// TIA Portal project "Energy_Drink_V15.1" (V15.1)

(* hardware
DEVICE "S7300/ET200M station_1"  S7-300 station
   slot 0: "Rail_0"  Rail  6ES7 390-1***0-0AA0
   slot 2: "ENERGY_DRINK_PROC"  CPU 314C-2 PN/DP  6ES7 314-6EH04-0AB0  V3.3
      slot 2: "PROFINET interface_1"  PN-IO
         slot 1: "Port_1"  Port
         slot 2: "Port_2"  Port
      slot 5: "DI 24/DO 16_1"  DI24/DO16
      slot 6: "AI 5/AO 2_1"  AI5/AO2
      slot 7: "Count_1"  Counter
      slot 8: "Positioning_1"  Positioning
   slot 4: "DI 16/DO 16x24VDC/0.5A_1"  DI16/DO16 x 24V / 0.5A  6ES7 323-1BL00-0AA0
   slot 5: "DI 8/DO 8x24VDC/0.5A_1"  DI8/DO8 x 24VDC / 0.5A  6ES7 323-1BH01-0AA0
   slot 6: "AI 2x12BIT_1"  AI2 x 12 bits  6ES7 331-7KB02-0AB0
   slot 7: "AO 4x12BIT_1"  AO4 x 12 bits  6ES7 332-5HD01-0AB0
DEVICE "HMI_1"  TP2200 Comfort
   slot 0: "HMI"  HMI  6AV2 124-0XC02-0AX0  13.0.1.0
   slot 1: "HMI_RT_1"  TP2200 Comfort  6AV2 124-0XC02-0AX0  13.0.1.0
   slot 5: "HMI_1.IE_CP_1"  Interfaz PROFINET
      slot 1: "Interfaz PROFINET_1"  Interfaz PROFINET
         slot 1: "Port_1"  Port
         slot 2: "Port_2"  Port
   slot 6: "HMI_1.IE_CP_2"  Interfaz PROFINET
      slot 1: "Interfaz PROFINET_GBit"  Interfaz PROFINET
         slot 1: "Port_1"  Port
   slot 7: "HMI_1.MPI/DP_CP_1"  Interfaz MPI/DP
*)

// ===== PLC "ENERGY_DRINK_PROC"  CPU 314C-2 PN/DP =====

VAR_GLOBAL   // PLC tag table "Default tag table"
   "M_Product_1" AT %MD100 : Real;
   "Tag_5" AT %MD50 : DWord;
   "Tag_6" AT %EW50 : Word;
   "Recipe_Num" AT %MW50 : Word;
   "M_Water_Flow" AT %MD112 : Real;
   "Num_Bach" AT %MW52 : Word;
   "Tag_3" AT %M10.0 : Bool;
   "Tag_7" AT %MD120 : Real;
   "Tag_13" AT %MD140 : Real;
   "M_Product_2" AT %MD104 : Real;
   "M_Product_3" AT %MD108 : Real;
   "M_Sirupe_Flow" AT %MD116 : Real;
   "FP_Conveyor_Act" AT %M255.7 : Bool;
   "FN_Bach_in_Prog" AT %M255.6 : Bool;
   "FN_TIMER.Q" AT %M255.5 : Bool;
   "FN_STOP_CMD" AT %M255.4 : Bool;
   "Tag_4" AT %MD200 : DWord;
   "Tag_10" AT %MW70 : Word;
   "Tag_11" AT %MD204 : DWord;
   "Tag_12" AT %M250.0 : Bool;
   "Tag_14" AT %M250.1 : Bool;
   "Tag_15" AT %MW60 : Int;
   "Tag_16" AT %MW62 : Int;
   "Tag_17" AT %MW64 : Int;
   "Tag_18" AT %MW66 : Int;
   "Tag_19" AT %MW68 : Int;
   "Tag_20" AT %MW72 : Int;
   "Tag_21" AT %MW74 : Int;
   "Tag_22" AT %MW76 : Int;
   "Tag_23" AT %MW78 : Int;
   "Tag_24" AT %MW80 : Int;
   "Tank1_Vlv" AT %AW800 : Word;
   "Tank2_Vlv" AT %AW802 : Word;
   "Tank3_Vlv" AT %AW804 : Word;
   "Sirupe_Vlv" AT %AW806 : Word;
   "Water_Vlv" AT %AW808 : Word;
   "Motor_VF" AT %AW810 : Word;
   "Tag_1" AT %MW82 : Int;
   "Tag_2" AT %M255.3 : Bool;
   "Tag_8" AT %M255.2 : Bool;
   "Tag_9" AT %M255.1 : Bool;
   "Tag_25" AT %M254.7 : Bool;
   "Tag_26" AT %M254.6 : Bool;
   "Tag_27" AT %M254.5 : Bool;
   "Total_Weight" AT %MD150 : Real;
   "Temp_Lim_Kg" AT %MD154 : Real;
   "Tag_29" AT %MD158 : Real;
   "Tag_28" AT %MD84 : DInt;
   "Tag_30" AT %M0.6 : Bool;
   "Tag_31" AT %M254.4 : Bool;
   "Tag_32" AT %M0.4 : Bool;
   "Tag_33" AT %M0.2 : Bool;
   "Tag_34" AT %M0.0 : Bool;
   "Tag_35" AT %M0.1 : Bool;
END_VAR

VAR_GLOBAL   // PLC tag table "VAR"
   "AUTO/MAN" AT %E0.0 : Bool;   // Switch Auto/Man
   "Start_Button" AT %E0.1 : Bool;   // Start switch "NO"
   "Stop_Button" AT %E0.2 : Bool;   // Stop switch "NC"
   "Emergency_Stop" AT %E0.3 : Bool;   // Emergency Stop "NC"
   "Man_Dis_Tk1_Vlv" AT %E136.1 : Bool;   // K1_Outlet gate Tank1 Switch
   "Man_Dis_Tk2_Vlv" AT %E136.2 : Bool;   // K2_Outlet gate Tank2 Switch
   "Man_Dis_Tk3_Vlv" AT %E136.3 : Bool;   // K3_Outlet gate Tank3 Switch
   "Man_Dis_Scale_Vlv" AT %E136.4 : Bool;   // K4_Outlet gate Scale Tank Switch
   "Convey_Man_Starter" AT %E136.5 : Bool;   // Starter start-delta motor Switch
   "Mixer_Man_Start" AT %E136.7 : Bool;   // VF Agitator motor Switch
   "Man_Dis_Mixer_Vlv" AT %E137.1 : Bool;   // K5_Outlet gate Mixer Tank Switch
   "Man_Water_Vlv" AT %E137.2 : Bool;   // K6_Water valve Switch
   "Man_Sirupe_Vlv" AT %E137.3 : Bool;   // K7_Sirupe valve Switch
   "Man_Fill_Tk1_Vlv" AT %E137.4 : Bool;   // K8_Filling valve Tank 1 Switch
   "Man_Fill_Tk2_Vlv" AT %E137.5 : Bool;   // K9_Filling valve Tank 2 Switch
   "Man_Fill_Tk3_Vlv" AT %E137.6 : Bool;   // K10_Filling valve Tank 3 Switch
   "OVL_Conveyor" AT %E137.7 : Bool;   // Overload Conveyor Motor
   "OVL_Mixer" AT %E138.0 : Bool;   // Overload VF Agitator
   "Recipe_1" AT %E138.1 : Bool;   // Recipe 1 Switch
   "Recipe_2" AT %E138.2 : Bool;   // Recipe 2 Switch
   "Recipe_3" AT %E138.3 : Bool;   // Recipe 3 Switch
   "Tank_1_Level" AT %EW800 : Int;
   "Tank_2_Level" AT %EW802 : Int;
   "Tank_3_Level" AT %EW804 : Int;
   "Weighing" AT %EW806 : Int;
   "Mixer_Tank_level" AT %EW808 : Int;
   "Water_Flow" AT %EW256 : Int;
   "Sirupe_Flow" AT %EW258 : Int;
   "Filling_Vlv_1_Opened" AT %E0.5 : Bool;
   "Filling_Vlv_1_Closed" AT %E0.6 : Bool;
   "Filling_Vlv_2_Closed" AT %E1.1 : Bool;
   "Filling_Vlv_2_Opened" AT %E1.2 : Bool;
   "Filling_Vlv_3_Closed" AT %E1.5 : Bool;
   "Filling_Vlv_3_Opened" AT %E1.6 : Bool;
   "Disch_Vlv_3_Opened" AT %E1.7 : Bool;
   "Disch_Vlv_3_Closed" AT %E2.0 : Bool;
   "Disch_Vlv_M_Opened" AT %E2.1 : Bool;
   "Disch_Vlv_M_Closed" AT %E2.2 : Bool;
   "Sirupe_Vlv_Closed" AT %E2.6 : Bool;
   "Disch_Vlv_1_Opened" AT %E0.7 : Bool;
   "Disch_Vlv_1_Closed" AT %E1.0 : Bool;
   "Disch_Vlv_2_Opened" AT %E1.3 : Bool;
   "Disch_Vlv_2_Closed" AT %E1.4 : Bool;
   "Water_Vlv_Closed" AT %E2.4 : Bool;
   "Water_Vlv_Opened" AT %E2.3 : Bool;
   "Sirupe_Vlv_Opened" AT %E2.5 : Bool;
   "Scale_Vlv_Opened" AT %E2.7 : Bool;
   "Scale_Vlv_Closed" AT %E136.0 : Bool;
   "Discharge_Vlv1" AT %A136.0 : Bool;   // Outlet gate Tank 1 rely
   "Discharge_Vlv2" AT %A136.1 : Bool;   // Outlet gate Tank 2 rely
   "Discharge_Vlv3" AT %A136.2 : Bool;   // Outlet gate Tank 3 rely
   "Scale_Dis_Vlv" AT %A136.3 : Bool;   // Outlet gate Scale Tank rely
   "Mixer_Dis_Vlv" AT %A136.4 : Bool;   // Outlet gate Mixer Tank rely
   "Filling_Vlv1" AT %A136.5 : Bool;   // Filling valve Tank 1 rely
   "Filling_Vlv2" AT %A136.6 : Bool;   // Filling valve Tank 2 rely
   "Filling_Vlv3" AT %A136.7 : Bool;   // Filling valve Tank 3 rely
   "Water_Vlv_Man" AT %A137.0 : Bool;
   "Sirupe_Vlv_Man" AT %A137.1 : Bool;
   "KM1_Main" AT %A137.2 : Bool;   // Conveyor Main Contactor
   "KM2_Star" AT %A137.3 : Bool;   // Conveyor Star Contactor
   "KM3_Delta" AT %A137.4 : Bool;
   "Mixer_Cleanning_Vlv" AT %A137.5 : Bool;   // Mixer Tank Cleaning valve
   "Start_Led" AT %A137.6 : Bool;   // Led Start
   "Stop_Led" AT %A137.7 : Bool;   // Led Stop
   "H3" AT %A0.0 : Bool;   // Led Emergency Stop
   "H4" AT %A0.1 : Bool;   // Led Conveyor Main Contactor
   "H5" AT %A0.2 : Bool;   // Led Conveyor Delta Contactor
   "H6" AT %A0.3 : Bool;   // Led aCELERATION VF Agitator
   "H7" AT %A0.4 : Bool;   // Led deceleration VF Agitator
   "H8" AT %A0.5 : Bool;   // Led Overload Conveyor
   "H9" AT %A0.6 : Bool;   // Led Overload VF Agitator
   "H10" AT %A0.7 : Bool;   // Led Conveyor Stopped
   "Reset_Button" AT %E0.4 : Bool;
   "Convey_Man_Stop" AT %E136.6 : Bool;
   "Mixer_Man_Stop" AT %E137.0 : Bool;
   "Enter_Selection" AT %E138.4 : Bool;
END_VAR

TYPE "UDT_RECIPE"
VERSION : 0.1
   STRUCT
      Recipe_Act : Bool;
      Num_Batches : Int;
      Product_1_Kg : Real;
      Product_2_Kg : Real;
      Product_3_Kg : Real;
      Water_Flow : Real;
      Sirupe_Flow : Real;
      Process_Time : Time;
   END_STRUCT;
END_TYPE

// folder: 01-MAIN PROCESS

DATA_BLOCK "Var_System_DB"   // DB1
{ S7_Optimized_Access := 'FALSE' }
VERSION : 0.1
   VAR
      Mixer_Motor : Struct
         Motor_Cmd : Bool;
         Man_Start : Bool;
         Man_Stop : Bool;
         Cmd_Start : Bool;
         Cmd_Stop : Bool;
         Overload : Bool;   // Memory activation Conveyor Motor Overload
         Led_Stopped : Bool;
         Led_Ovl : Bool;   // Memory activation Led Conveyor Motor Overload
         Acel_Led : Bool;
         Decel_Led : Bool;
         Feedback : Bool;
         FP_Start : Bool;
         FP_Timer : Bool;
         FN_Stop : Bool;
         State : Bool;
         Aceleration_T : Time := T#10S;
         Deceleration_T : Time := T#6S;
         PV : Int;
      END_STRUCT;
      System_Generic : Struct
         "Auto/Man" : Bool;
         Man_Mode : Bool;
         Start : Bool;
         Stop : Bool;
         Enter_Selection : Bool;
         Emergency_Stop : Bool;
         Man_Start_Process : Bool;
         Stop_Process : Bool;
         System_Act : Bool := false;   // System Active
         System_Failure : Bool;   // System Failure
         System_Alarm : Bool;   // System Alarm
         No_Process : Bool;
         Bach_In_Progress : Bool;
         Conveyor_Station : Bool;
         Mixer_Station : Bool;
         T_Mixer_Station : Bool;
         Always_True : Bool := true;
         Always_False : Bool;
         Recipe_num : Word;
         "HMI/OPERATOR" : Int;
      END_STRUCT;
      Conveyor_Belt : Struct
         Motor_Cmd : Bool;
         Man_Start : Bool;
         Man_Stop : Bool;
         M_Stop : Bool;
         M_Main : Bool;   // Memory activation Main Contactor
         M_Star : Bool;   // Memory activation Star Contactor
         M_Delta : Bool;   // Memory activation Delta Contactor
         M_Overload : Bool;   // Memory activation Conveyor Motor Overload
         M_Led_Main : Bool;   // Memory activation Led Main Contactor
         M_Led_Delta : Bool;   // Memory activation Led Delta Contactor
         M_Led_Stop : Bool;
         M_Led_Ovl : Bool;   // Memory activation Led Conveyor Motor Overload
         M_Feedback : Bool;
         Timer_Act : Bool;
         State : Bool;
         Move_Counter : Bool;
         Move_Increment : Int;
         T_Star : Time := T#6S;
         Time_Conveyor_Act : Time := T#12S;
      END_STRUCT;
      Sirupe_Flow_Meter : Struct
         Ret_Val : Word;
         Flow_Meter : Int;
         Flow_PV : Real;   // Liters per second
         Low_Lim : Real;
         High_Lim : Real;
      END_STRUCT;
      Sirupe_Valve : Struct
         Vlv_Cmd : Bool;
         Vlv_Opened : Bool;
         Vlv_Closed : Bool;
         Vlv_Open_Cmd : Bool;
         Vlv_Feedback : Bool;
         FP_Reset : Bool;
         Ret_Value : Word;
         Vlv_Actuator_Cmd : Int;
         "%_Vlv_Opened" : DInt;
         Increment_T : Time := T#0MS;
      END_STRUCT;
      Tk101 : Struct
         Vlv_Cmd : Bool;
         Vlv_Opened : Bool;
         Vlv_Closed : Bool;
         Vlv_Feedback : Bool;
         Low_Level_Alarm : Bool;
         High_Level_Alarm : Bool;
         Vlv_Alarm : Bool;
         Vlv_Open_Cmd : Bool;
         Vlv_Close_Cmd : Bool;
         Ret_Value : Word;
         Vlv_Actuator_Cmd : Int;
         Double_Feedback : Int := 3;
         Inverse : Int := 4;
         LT_Value : Int;   // Level Transmitter
         "%_Vlv_Opened" : DInt;
         "Level_%" : DInt;
         Level_Liters : Real;
         Min_level : Real := 15.0;
         Max_level : Real := 90.0;
         Radius : Real := 1.5;
         Height : Real := 10.0;
         Scale_Kg : Real;
      END_STRUCT;
      TK101_FILLING_VLV : Struct
         Vlv_Cmd : Bool;
         Vlv_Opened : Bool;
         Vlv_Closed : Bool;
         Vlv_Feedback : Bool;
         Open_Vlv_Cmd : Bool;
         Close_Vlv_Cmd : Bool;
         Single_Actuation : Int := 1;
         Double_Feedback : Int := 3;
      END_STRUCT;
      Tk102 : Struct
         Vlv_Cmd : Bool;
         Vlv_Opened : Bool;
         Vlv_Closed : Bool;
         Vlv_Feedback : Bool;
         Low_Level_Alarm : Bool;
         High_Level_Alarm : Bool;
         Vlv_Alarm : Bool;
         Vlv_Open_Cmd : Bool;
         Vlv_Close_Cmd : Bool;
         Ret_Value : Word;
         Vlv_Actuator_Cmd : Int;
         Double_Feedback : Int := 3;
         Inverse : Int := 4;
         LT_Value : Int;
         "%_Vlv_Opened" : DInt;
         "Level_%" : DInt;
         Level_Liters : Real;
         Min_level : Real := 15.0;
         Max_level : Real := 90.0;
         Radius : Real := 1.5;
         Height : Real := 10.0;
         Scale_Kg : Real;
      END_STRUCT;
      TK102_FILLING_VLV : Struct
         Vlv_Cmd : Bool;
         Vlv_Opened : Bool;
         Vlv_Closed : Bool;
         Vlv_Feedback : Bool;
         Open_Vlv_Cmd : Bool;
         Close_Vlv_Cmd : Bool;
         Single_Actuation : Int := 1;
         Double_Feedback : Int := 3;
      END_STRUCT;
      Tk103 : Struct
         Vlv_Cmd : Bool;
         Vlv_Opened : Bool;
         Vlv_Closed : Bool;
         Vlv_Feedback : Bool;
         Low_Level_Alarm : Bool;
         High_Level_Alarm : Bool;
         Vlv_Alarm : Bool;
         Vlv_Open_Cmd : Bool;
         Vlv_Close_Cmd : Bool;
         Ret_Value : Word;
         Vlv_Actuator_Cmd : Int;
         Double_Feedback : Int := 3;
         Inverse : Int := 4;
         LT_Value : Int;
         "%_Vlv_Opened" : DInt;
         "Level_%" : DInt;
         Level_Liters : Real;
         Min_level : Real := 15.0;
         Max_level : Real := 90.0;
         Radius : Real := 1.5;
         Height : Real := 10.0;
         Scale_Kg : Real;
      END_STRUCT;
      TK103_FILLING_VLV : Struct
         Vlv_Cmd : Bool;
         Vlv_Opened : Bool;
         Vlv_Closed : Bool;
         Vlv_Feedback : Bool;
         Open_Vlv_Cmd : Bool;
         Close_Vlv_Cmd : Bool;
         Single_Actuation : Int := 1;
         Double_Feedback : Int := 3;
      END_STRUCT;
      Tk104_MIXER : Struct
         Tank_Cmd : Bool;
         Dis_Vlv_Cmd : Bool := false;
         Vlv_Opened : Bool;
         Vlv_Closed : Bool;
         Open_Vlv_Cmd : Bool;
         Close_Vlv_Cmd : Bool;
         Single_Actuation : Int := 1;
         Double_Feedback : Int := 3;
         Vlv_Feedback : Bool;
         Low_Level_Alarm : Bool;
         High_Level_Alarm : Bool;
         Vlv_Alarm : Bool;
         FN_Agitator : Bool;
         Ret_Value : Word;
         Vlv_Actuator_Cmd : Int;
         Proportional_Feedback : Int := 4;
         Inverse_Mode : Int := 5;
         LT_Value : Int;
         "%_Vlv_Opened" : DInt;
         "Level_%" : DInt;
         Level_Liters : Real;
         Min_level : Real := 1.5;
         Max_level : Real := 9.0;
         Radius : Real := 1.5;
         Height : Real := 10.0;
         Scale_Kg : Real;
      END_STRUCT;
      Water_Flow_Meter : Struct
         Ret_Val : Word;
         Flow_Meter : Int;
         Flow_PV : Real;   // Liters per second
         Low_Lim : Real;
         High_Lim : Real := 15.0;
      END_STRUCT;
      Water_Valve : Struct
         Vlv_Cmd : Bool;
         Vlv_Opened : Bool;
         Vlv_Closed : Bool;
         Vlv_Open_Cmd : Bool;
         Vlv_Feedback : Bool;
         Vlv_Alarm : Bool;
         FP_Start : Bool;
         FP_Stop : Bool;
         Vlv_Act : Bool;
         Ret_Value : Word;
         Vlv_Actuator_Cmd : Int;
         Proportional_Feedback : Int := 4;
         Proportional_Mode : Int := 3;
         "%_Vlv_Opened" : DInt;
         PV : Real := 50.0;
      END_STRUCT;
      Weighing_Process : Struct
         Weighing_In_Progress : Bool;
         Weighing_Value : Int;
         State : Int := 0;
         Max_Kg : Real := 100000.0;
         Min_Kg : Real;
         PV : Real;   // Process Value
      END_STRUCT;
      Scale_Discharge_Vlv : Struct
         Vlv_Cmd : Bool;
         Vlv_Opened : Bool;
         Vlv_Closed : Bool;
         Vlv_Feedback : Bool;
         Open_Vlv : Bool;
         Open_Vlv_Cmd : Bool;
         Single_Actuation : Int := 1;
         Double_Feedback : Int := 3;
      END_STRUCT;
      Cleanning_Process : Struct
         Vlv_Open_Cmd : Bool;
      END_STRUCT;
   END_VAR
BEGIN
END_DATA_BLOCK

DATA_BLOCK "HMI_VAR"   // DB20
{ S7_Optimized_Access := 'FALSE' }
VERSION : 0.1
   VAR
      Recipe_Selection : Array[1..4] of Bool;   // Diferent types of recipes
      Test_Recipe : Struct
         Products : Array[1..3] of Real;
         Flows : Array[1..2] of Real;
      END_STRUCT;
      Warnings : Word;
      Man_Valves : Struct
         Filling_Vlv1 : Bool;
         Filling_Vlv2 : Bool;
         Filling_Vlv3 : Bool;
         Scale_Vlv : Bool;
         Mixer_Discharge_Vlv : Bool;
         Discharge_Vlv1 : Bool;
         Discharge_Vlv2 : Bool;
         Discharge_Vlv3 : Bool;
         Water_Vlv : Bool;
         Sirupe_Vlv : Bool;
      END_STRUCT;
      Man_Motors : Struct
         Start_Conveyor : Bool;
         Stop_Conveyor : Bool;
         Start_Mixer : Bool;
         Stop_Mixer : Bool;
      END_STRUCT;
      Conveyor : Struct
         Belt : Bool;
         Container_Move : Int;
      END_STRUCT;
      Mixer : Struct
         Agitator_1 : Bool;
         Agitator_2 : Bool;
      END_STRUCT;
      Act_System : Bool;
      Stop_System : Bool := true;
      "Auto/Manual" : Bool;
      Enter_Selection : Bool;
      Start_Process : Bool;
      Reset_Selection : Bool;
   END_VAR
BEGIN
   Test_Recipe.Products[1] := 0.0;
END_DATA_BLOCK

// folder: 03-TANK MANAGEMENT

DATA_BLOCK "TK101_DISCHARGE_VLV_DB"   // DB2
{ S7_Optimized_Access := 'FALSE' }
VERSION : 0.1
// stored: InstanceOfName GENERIC_VALVE
"GENERIC_VALVE"
BEGIN
END_DATA_BLOCK

DATA_BLOCK "TK101_FILLING_VLV_DB"   // DB3
{ S7_Optimized_Access := 'FALSE' }
VERSION : 0.1
// stored: InstanceOfName GENERIC_VALVE
"GENERIC_VALVE"
BEGIN
END_DATA_BLOCK

DATA_BLOCK "TK102_FILLING_VLV_DB"   // DB4
{ S7_Optimized_Access := 'FALSE' }
VERSION : 0.1
// stored: InstanceOfName GENERIC_VALVE
"GENERIC_VALVE"
BEGIN
END_DATA_BLOCK

DATA_BLOCK "TK102_DISCHARGE_VLV_DB"   // DB5
{ S7_Optimized_Access := 'FALSE' }
VERSION : 0.1
// stored: InstanceOfName GENERIC_VALVE
"GENERIC_VALVE"
BEGIN
END_DATA_BLOCK

DATA_BLOCK "TK103_FILLING_VLV_DB"   // DB6
{ S7_Optimized_Access := 'FALSE' }
VERSION : 0.1
// stored: InstanceOfName GENERIC_VALVE
"GENERIC_VALVE"
BEGIN
END_DATA_BLOCK

DATA_BLOCK "TK103_DISCHARGE_VLV_DB"   // DB7
{ S7_Optimized_Access := 'FALSE' }
VERSION : 0.1
// stored: InstanceOfName GENERIC_VALVE
"GENERIC_VALVE"
BEGIN
END_DATA_BLOCK

// folder: 04-OPERATOR MANAGEMENT

DATA_BLOCK "RECIPE_1_DB"   // DB10
{ S7_Optimized_Access := 'FALSE' }
VERSION : 0.1
   VAR
      Recipe1 : "UDT_RECIPE";
   END_VAR
BEGIN
   Recipe1.Product_1_Kg := 30000.0;
   Recipe1.Product_2_Kg := 25000.0;
   Recipe1.Product_3_Kg := 15000.0;
   Recipe1.Water_Flow := 7.5;
   Recipe1.Sirupe_Flow := 2.5;
END_DATA_BLOCK

DATA_BLOCK "RECIPE_2_DB"   // DB11
{ S7_Optimized_Access := 'FALSE' }
VERSION : 0.1
   VAR
      Recipe2 : "UDT_RECIPE";
   END_VAR
BEGIN
   Recipe2.Product_1_Kg := 35000.0;
   Recipe2.Product_2_Kg := 22500.0;
   Recipe2.Product_3_Kg := 17850.0;
   Recipe2.Water_Flow := 7.5;
   Recipe2.Sirupe_Flow := 3.3;
END_DATA_BLOCK

DATA_BLOCK "RECIPE_3_DB"   // DB12
{ S7_Optimized_Access := 'FALSE' }
VERSION : 0.1
   VAR
      Recipe3 : "UDT_RECIPE";
   END_VAR
BEGIN
   Recipe3.Product_1_Kg := 12500.0;
   Recipe3.Product_2_Kg := 9000.0;
   Recipe3.Product_3_Kg := 8525.0;
   Recipe3.Water_Flow := 7.2;
   Recipe3.Sirupe_Flow := 3.7;
END_DATA_BLOCK

DATA_BLOCK "TEST_RECIPE_DB"   // DB13
{ S7_Optimized_Access := 'FALSE' }
VERSION : 0.1
   VAR
      Test : "UDT_RECIPE";
   END_VAR
BEGIN
END_DATA_BLOCK

DATA_BLOCK "SCALE_DISCHARGE_VLV_DB"   // DB15
{ S7_Optimized_Access := 'FALSE' }
VERSION : 0.1
// stored: InstanceOfName GENERIC_VALVE
"GENERIC_VALVE"
BEGIN
END_DATA_BLOCK

// folder: 05-CONVEYOR MANAGEMENT

DATA_BLOCK "CONVEYOR_DB"   // DB14
{ S7_Optimized_Access := 'FALSE' }
VERSION : 0.1
// stored: InstanceOfName STAR/DELTA_STARTER
"STAR/DELTA_STARTER"
BEGIN
END_DATA_BLOCK

// folder: 06-MIXER MANAGEMENT

DATA_BLOCK "WATER_VALVE_DB"   // DB8
{ S7_Optimized_Access := 'FALSE' }
VERSION : 0.1
// stored: InstanceOfName GENERIC_VALVE
"GENERIC_VALVE"
BEGIN
END_DATA_BLOCK

DATA_BLOCK "INCREMENTAL_PULSE_VLV_DB"   // DB9
{ S7_Optimized_Access := 'FALSE' }
VERSION : 0.1
// stored: InstanceOfName INCREMENTAL_PULSE_VLV
"INCREMENTAL_PULSE_VLV"
BEGIN
END_DATA_BLOCK

DATA_BLOCK "MIXER_DISCHARGE_VLV"   // DB17
{ S7_Optimized_Access := 'FALSE' }
VERSION : 0.1
// stored: InstanceOfName GENERIC_VALVE
"GENERIC_VALVE"
BEGIN
END_DATA_BLOCK

DATA_BLOCK "MIXER_MOTOR_DB"   // DB18
{ S7_Optimized_Access := 'FALSE' }
VERSION : 0.1
// stored: InstanceOfName MOTOR_ACELERATION_RAMP
"MOTOR_ACELERATION_RAMP"
BEGIN
END_DATA_BLOCK

// folder: 01-MAIN PROCESS

FUNCTION "HMI_CONTROL" : Void   // FC2, STL
{ S7_Optimized_Access := 'FALSE' }
VERSION : 0.1
BEGIN

REGION Network 1: /************************MOVE DATA FROM HMI TO DB*****************************************/
   // MOVE THE DATA INTRODUCED IN HMI TO RECIPE TEST DB
   // WITH THIS INSTRUCTION WE MOVE THE PRODUCT AND FLOWS DATA
   // TO SET UP A RECIPE TEST ENVIROMENT.

         CALL  BLKMOV
         ( SRCBLK  := P#DB20.DBX2.0 BYTE 20,
           RET_VAL := "Tag_1",
           DSTBLK  := P#DB13.DBX4.0 BYTE 20
         );
END_REGION

REGION Network 2: /************************HMI WARNINGS*****************************************/
   //********************OVERLOAD WARNINGS***********************************//

   // CONVEYOR OVERLOAD WARNING
         AN    "Var_System_DB".Conveyor_Belt.M_Overload;
         =     %DB20.DBX22.0;

   // MIXER OVERLOAD WARNING
         AN    "Var_System_DB".Mixer_Motor.Overload;
         =     %DB20.DBX22.1;


   //********************TANKS WARNINGS AND ALARMS***********************************//

   // TANK 1 LOW LEVEL
         A     "Var_System_DB".Tk101.Low_Level_Alarm;
         =     %DB20.DBX22.2;

         A     "Var_System_DB".Tk101.High_Level_Alarm;
         =     %DB20.DBX22.3;

   // TANK 2 LOW LEVEL
         A     "Var_System_DB".Tk102.Low_Level_Alarm;
         =     %DB20.DBX22.4;

         A     "Var_System_DB".Tk102.High_Level_Alarm;
         =     %DB20.DBX22.5;


   // TANK 3 LOW LEVEL
         A     "Var_System_DB".Tk103.Low_Level_Alarm;
         =     %DB20.DBX22.6;

         A     "Var_System_DB".Tk103.High_Level_Alarm;
         =     %DB20.DBX22.7;
END_REGION

REGION Network 3: /************************MANUAL MODE*****************************************/
   //********************************MANUAL MODE ACTIVE*************************************//

   // IF AUTO MODE = 1
         A     "Var_System_DB".System_Generic.Man_Mode;
         JCN   _1001;

   //********************************FILLING VALVES*************************************//
   // MAN FILLING VALVE 1
         A     "HMI_VAR".Man_Valves.Filling_Vlv1;
         =     "Var_System_DB".TK101_FILLING_VLV.Open_Vlv_Cmd;

   // MAN FILLING VALVE 2
         A     "HMI_VAR".Man_Valves.Filling_Vlv2;
         =     "Var_System_DB".TK102_FILLING_VLV.Open_Vlv_Cmd;

   // MAN FILLING VALVE 3
         A     "HMI_VAR".Man_Valves.Filling_Vlv3;
         =     "Var_System_DB".TK103_FILLING_VLV.Open_Vlv_Cmd;

   //********************************DISCHARGE VALVES*************************************//

   // DISCHARGE VALVE 1
         A     "HMI_VAR".Man_Valves.Discharge_Vlv1;
         JCN   _1002;
         L     27648;
         T     "Var_System_DB".Weighing_Process.PV;
   _1002:NOP   0;

   // DISCHARGE VALVE 2
         A     "HMI_VAR".Man_Valves.Discharge_Vlv2;
         JCN   _1003;
         L     27648;
         T     "Var_System_DB".Weighing_Process.PV;
   _1003:NOP   0;

   // DISCHARGE VALVE 3
         A     "HMI_VAR".Man_Valves.Discharge_Vlv3;
         JCN   _1004;
         L     27648;
         T     "Var_System_DB".Weighing_Process.PV;
   _1004:NOP   0;

   //********************************MIXER STATION*************************************//

   // MIXER MOTOR
         A     "HMI_VAR".Man_Motors.Start_Mixer;
         =     "Var_System_DB".Mixer_Motor.Motor_Cmd;

   // WATER VALVE
         A     "HMI_VAR".Man_Valves.Water_Vlv;
         JCN   _1005;
         L     10.0;
         T     "M_Water_Flow";
   _1005:NOP   0;

   // WATER VALVE
         A     "HMI_VAR".Man_Valves.Sirupe_Vlv;
         JCN   _1006;
         L     27648;
         T     "Var_System_DB".Sirupe_Valve.Vlv_Actuator_Cmd;
   _1006:NOP   0;

   _1001:NOP   0;
END_REGION

REGION Network 4: /************************AGITATOR MOVEMENT*****************************************/
         A     "Var_System_DB".Mixer_Motor.Feedback;
         A     "Tag_32";
         =     "HMI_VAR".Mixer.Agitator_1;
END_REGION

REGION Network 5: /************************CONVEYOR MOVEMENT*****************************************/
         A     "Var_System_DB".Conveyor_Belt.M_Feedback;
         A     "Tag_33";
         FP    "Tag_31";
         JCN   _1010;
         L     2;
         L     "HMI_VAR".Conveyor.Container_Move;
         +I;
         T     "HMI_VAR".Conveyor.Container_Move;

         A(;
         L     "HMI_VAR".Conveyor.Container_Move;
         L     100;
         ==I;
         );
         JCN   _1011;
         L     0;
         T     "HMI_VAR".Conveyor.Container_Move;
   _1011:NOP   0;


   _1010:NOP   0;
END_REGION
END_FUNCTION

FUNCTION "TANK_LEVEL" : Void   // FC8, STL
{ S7_Optimized_Access := 'FALSE' }
VERSION : 0.1
   VAR_INPUT
      Tank_Cmd : Bool;
      LT_Value : Int;   // Level transmiter value
      Radius : Real;   // Tank radius
      Height : Real;   // Tank height
      Low_Level : Real;
      High_Level : Real;
   END_VAR
   VAR_OUTPUT
      High_Alarm : Bool;
      Low_Alarm : Bool;
      Level_Liters : Real;   // Tank level in liters
      Ret_Value : Word;
   END_VAR
   VAR_IN_OUT
      "Level_%" : DInt;   // Tank level in %
   END_VAR
   VAR_TEMP
      Temp_Level : Real;
   END_VAR
BEGIN

REGION Network 1: *****************************SENSOR SCALING MANAGEMENT*************************************
   // LEVEL SENSOR SCALING FROM OUT SIGNAL
         CALL  SCALE
         ( IN      := #LT_Value,
           HI_LIM  := #Height,
           LO_LIM  := 0.0,
           BIPOLAR := FALSE,
           RET_VAL := #Ret_Value,
           OUT     := #Temp_Level
         );

   // MAP VAR TEMP_LEVEL TO LEVEL_% TO VISUALIZE THE LEVEL OF THE TANK
         L     #Temp_Level;
         L     10.0;
         *R;
         RND;
         T     #"Level_%";  // LEVEL IN %
END_REGION

REGION Network 2: *******************************CALCULATE VOLUME TANK IN LITERS****************************
   // IF TANK COMMAND => CALCULATE VOLUME IN LITERS BASED ON INPUT PARAMETERS
         A     #Tank_Cmd;
         JCN   _001;
         L     #Radius;
         SQR;
         L     3.1416;
         *R;
         L     #Temp_Level;
         *R;
         L     1000.0;
         *R;
         T     #Level_Liters;  // LEVEL IN LITERS

   _001: NOP   0;
END_REGION

REGION Network 3: ********************************HIGH LEVEL ALARM**********************************************
   // IF LEVEL >= HIGH_LEVEL => SET HIGH ALARM
         A     #Tank_Cmd;
         A(;
         L     #"Level_%";
         DTR;
         L     #High_Level;
         >=R;
         );
         =     #High_Alarm;
END_REGION

REGION Network 4: ********************************LOW LEVEL ALARM**********************************************
   // IF LEVEL <= LOW_LEVEL => SET HIGH ALARM
         A     #Tank_Cmd;
         A(;
         L     #"Level_%";
         DTR;
         L     #Low_Level;
         <=R;
         );
         =     #Low_Alarm;
END_REGION
END_FUNCTION

FUNCTION "PROCESS_CONTROL" : Void   // FC14, FBD
{ S7_Optimized_Access := 'FALSE' }
VERSION : 0.1
BEGIN

REGION Network 1: ***************************** TANKS MANAGEMENT********************************************/
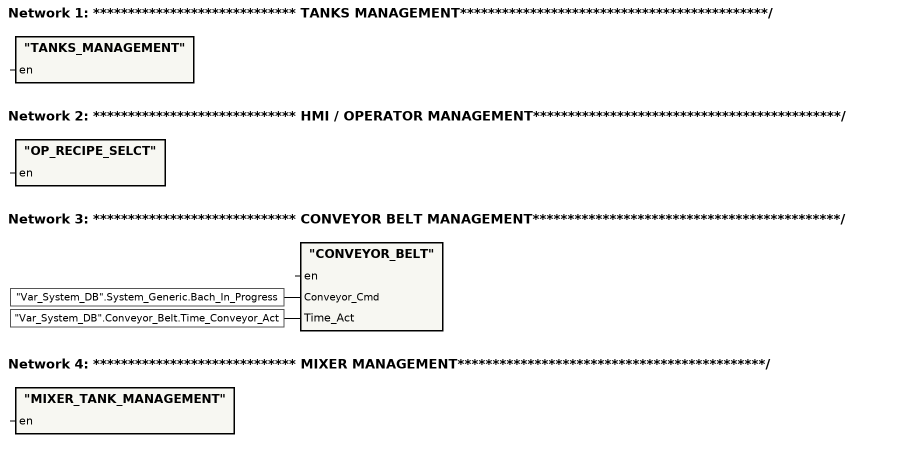
   "TANKS_MANAGEMENT"();
END_REGION

REGION Network 2: ***************************** HMI / OPERATOR MANAGEMENT********************************************/
   "OP_RECIPE_SELCT"();
END_REGION

REGION Network 3: ***************************** CONVEYOR BELT MANAGEMENT********************************************/
   "CONVEYOR_BELT"(Conveyor_Cmd := "Var_System_DB".System_Generic.Bach_In_Progress,
                   Time_Act := "Var_System_DB".Conveyor_Belt.Time_Conveyor_Act);
END_REGION

REGION Network 4: ***************************** MIXER MANAGEMENT********************************************/
   "MIXER_TANK_MANAGEMENT"();
END_REGION
END_FUNCTION

ORGANIZATION_BLOCK "Main"   // OB1, FBD
TITLE = "Main Program Sweep (Cycle)"
{ S7_Optimized_Access := 'FALSE' }
VERSION : 0.1
   VAR_TEMP
      OB1_EV_CLASS : Byte;   // Bits 0-3 = 1 (Coming event), Bits 4-7 = 1 (Event class 1)
      OB1_SCAN_1 : Byte;   // 1 (Cold restart scan 1 of OB 1), 3 (Scan 2-n of OB 1)
      OB1_PRIORITY : Byte;   // Priority of OB Execution
      OB1_OB_NUMBR : Byte;   // 1 (Organization block 1, OB1)
      OB1_RESERVED_1 : Byte;   // Reserved for system
      OB1_RESERVED_2 : Byte;   // Reserved for system
      OB1_PREV_CYCLE : Int;   // Cycle time of previous OB1 scan (milliseconds)
      OB1_MIN_CYCLE : Int;   // Minimum cycle time of OB1 (milliseconds)
      OB1_MAX_CYCLE : Int;   // Maximum cycle time of OB1 (milliseconds)
      OB1_DATE_TIME : Date_And_Time;   // Date and time OB1 started
   END_VAR
BEGIN

REGION Network 1: *********************** SENSOR AND ACTUATORS MANAGEMENT********************************************/
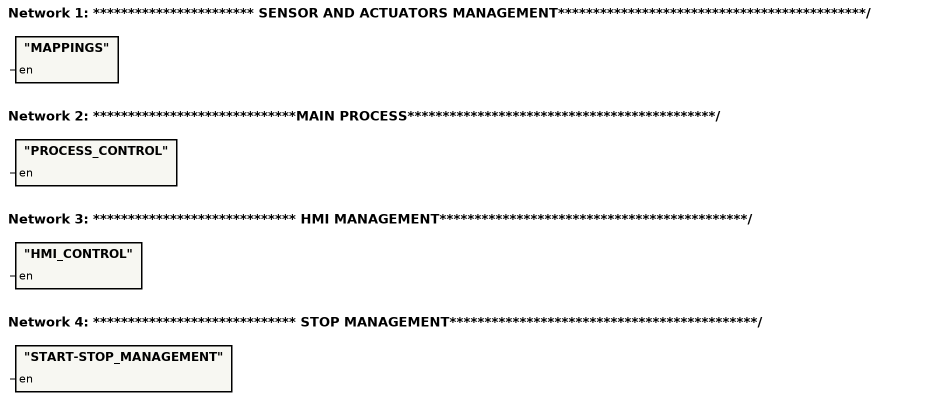
   "MAPPINGS"();
END_REGION

REGION Network 2: *****************************MAIN PROCESS********************************************/
   "PROCESS_CONTROL"();
END_REGION

REGION Network 3: ***************************** HMI MANAGEMENT********************************************/
   "HMI_CONTROL"();
END_REGION

REGION Network 4: ***************************** STOP MANAGEMENT********************************************/
   "START-STOP_MANAGEMENT"();
END_REGION
END_ORGANIZATION_BLOCK

// folder: 01-MAIN PROCESS/SENSORS ACTUATORS MANAGEMENT

FUNCTION "MAPPINGS" : Void   // FC15, FBD
{ S7_Optimized_Access := 'FALSE' }
VERSION : 0.1
BEGIN

REGION Network 1: ***************************** ACTUATORS MAPPING ********************************************/
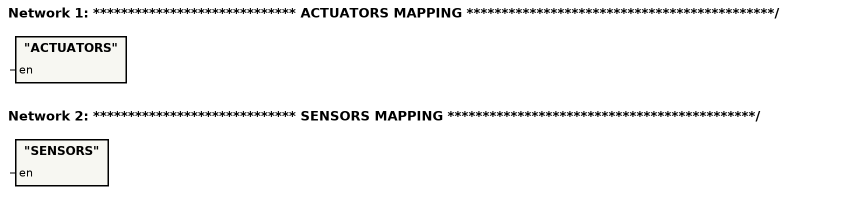
   "ACTUATORS"();
END_REGION

REGION Network 2: ***************************** SENSORS MAPPING ********************************************/
   "SENSORS"();
END_REGION
END_FUNCTION

FUNCTION "SENSORS" : Void   // FC18, STL
{ S7_Optimized_Access := 'FALSE' }
VERSION : 0.1
BEGIN

REGION Network 1: *****************************TANK 1 MAPPINGS*************************************
   // TANK LEVEL 1
         L     "Tank_1_Level":P;
         T     "Var_System_DB".Tk101.LT_Value;

   // FILLING VALVE
         A     "Filling_Vlv_1_Closed";
         =     "Var_System_DB".TK101_FILLING_VLV.Vlv_Closed;

         A     "Filling_Vlv_1_Opened";
         =     "Var_System_DB".TK101_FILLING_VLV.Vlv_Opened;

         A     "Man_Fill_Tk1_Vlv";
         =     "Var_System_DB".TK101_FILLING_VLV.Open_Vlv_Cmd;

   // DISCHARGE VALVE
         A     "Disch_Vlv_1_Closed";
         =     "Var_System_DB".Tk101.Vlv_Closed;

         A     "Disch_Vlv_1_Opened";
         =     "Var_System_DB".Tk101.Vlv_Opened;
END_REGION

REGION Network 2: *****************************TANK 2 MAPPINGS*************************************
   // TANK LEVEL 2
         L     "Tank_2_Level":P;
         T     "Var_System_DB".Tk102.LT_Value;

   // FILLING VALVE
         A     "Filling_Vlv_2_Closed";
         =     "Var_System_DB".TK102_FILLING_VLV.Vlv_Closed;

         A     "Filling_Vlv_2_Opened";
         =     "Var_System_DB".TK102_FILLING_VLV.Vlv_Opened;

         A     "Man_Fill_Tk2_Vlv";
         =     "Var_System_DB".TK102_FILLING_VLV.Open_Vlv_Cmd;

   // DISCHARGE VALVE
         A     "Disch_Vlv_2_Closed";
         =     "Var_System_DB".Tk102.Vlv_Closed;

         A     "Disch_Vlv_2_Opened";
         =     "Var_System_DB".Tk102.Vlv_Opened;
END_REGION

REGION Network 3: *****************************TANK 3 MAPPINGS*************************************
   // TANK LEVEL 3
         L     "Tank_3_Level":P;
         T     "Var_System_DB".Tk103.LT_Value;

   // FILLING VALVE
         A     "Filling_Vlv_3_Closed";
         =     "Var_System_DB".TK103_FILLING_VLV.Vlv_Closed;

         A     "Filling_Vlv_3_Opened";
         =     "Var_System_DB".TK103_FILLING_VLV.Vlv_Opened;

         A     "Man_Fill_Tk3_Vlv";
         =     "Var_System_DB".TK103_FILLING_VLV.Open_Vlv_Cmd;
   // DISCHARGE VALVE
         A     "Disch_Vlv_3_Closed";
         =     "Var_System_DB".Tk103.Vlv_Closed;

         A     "Disch_Vlv_3_Opened";
         =     "Var_System_DB".Tk103.Vlv_Opened;
END_REGION

REGION Network 4: *****************************MIXER TANK MAPPINGS*************************************
   // MIXER TANK LEVEL
         L     "Mixer_Tank_level":P;
         T     "Var_System_DB".Tk104_MIXER.LT_Value;

   // WATER FLOW METER
         L     "Water_Flow":P;
         T     "Var_System_DB".Water_Flow_Meter.Flow_Meter;

   // WATER VALVE
         A     "Water_Vlv_Closed";
         =     "Var_System_DB".Water_Valve.Vlv_Closed;

         A     "Water_Vlv_Opened";
         =     "Var_System_DB".Water_Valve.Vlv_Opened;

   // SIRUPE FLOW METER
         L     "Sirupe_Flow":P;
         T     "Var_System_DB".Sirupe_Flow_Meter.Flow_Meter;

   // SIRUPE VALVE
         A     "Sirupe_Vlv_Closed";
         =     "Var_System_DB".Sirupe_Valve.Vlv_Closed;

         A     "Sirupe_Vlv_Opened";
         =     "Var_System_DB".Sirupe_Valve.Vlv_Opened;

   // DISCHARGE VALVE
         A     "Disch_Vlv_M_Closed";
         =     "Var_System_DB".Tk104_MIXER.Vlv_Closed;

         A     "Disch_Vlv_M_Opened";
         =     "Var_System_DB".Tk104_MIXER.Vlv_Opened;
END_REGION

REGION Network 5: *****************************SCALE*************************************
   // SCALE SENSOR
         L     "Weighing":P;
         T     "Var_System_DB".Weighing_Process.Weighing_Value;

   // DISCHARGE VALVE
         A     "Scale_Vlv_Closed";
         =     "Var_System_DB".Scale_Discharge_Vlv.Vlv_Closed;

         A     "Scale_Vlv_Opened";
         =     "Var_System_DB".Scale_Discharge_Vlv.Vlv_Opened;
END_REGION

REGION Network 6: *****************************CONVEYOR*************************************
   // CONVEYOR MOTOR MANUAL START
         A     "Convey_Man_Starter";
         O     "HMI_VAR".Man_Motors.Start_Conveyor;
         =     "Var_System_DB".Conveyor_Belt.Man_Start;

   // CONVEYOR MOTOR MANUAL STOP
         A     "Convey_Man_Stop";
         =     "Var_System_DB".Conveyor_Belt.Man_Stop;

   // CONVEYOR MOTOR OVERLOAD
         A     "OVL_Conveyor";
         =     "Var_System_DB".Conveyor_Belt.M_Overload;
END_REGION

REGION Network 7: *****************************MIXER MOTOR VF*************************************
   // MIXER MANUAL MOTOR START
         A     "Mixer_Man_Start";
         O     "HMI_VAR".Man_Motors.Start_Mixer;
         =     "Var_System_DB".Mixer_Motor.Man_Start;

   // MIXER MANUAL MOTOR STOP
         A     "Mixer_Man_Stop";
         =     "Var_System_DB".Mixer_Motor.Man_Stop;

   // MIXER MOTOR OVERLOAD
         A     "OVL_Mixer";
         =     "Var_System_DB".Mixer_Motor.Overload;
END_REGION

REGION Network 8: *****************************SIRUPE AND WATER VALVE*************************************
   // SIRUPE VALVE
         A     "Sirupe_Vlv_Man";
         =     "Var_System_DB".Sirupe_Valve.Vlv_Open_Cmd;

   // WATER VALVE
         A     "Water_Vlv_Man";
         =     "Var_System_DB".Water_Valve.Vlv_Open_Cmd;
END_REGION

REGION Network 9: *****************************AUTO/MANUAL*************************************
   // AUTO = 0 / MANUAL = 1
         A     "AUTO/MAN";
         O     "HMI_VAR"."Auto/Manual";
         =     "Var_System_DB".System_Generic."Auto/Man";

   // ENTER RECIPE SELECTION
         A     "Enter_Selection";
         =     "Var_System_DB".System_Generic.Enter_Selection;
END_REGION
END_FUNCTION

FUNCTION "ACTUATORS" : Void   // FC19, STL
TITLE = ************FUNCTION TO MAP THE PROCESS ACTUATORS TO ITS CORRESPONDING VAR********************************************/
{ S7_Optimized_Access := 'FALSE' }
VERSION : 0.1
BEGIN

REGION Network 1: *****************************ANALOG ACTUATORS********************************************/
   // TANK 1 DISCHARGE VALVE
         L     "Var_System_DB".Tk101.Vlv_Actuator_Cmd;
         T     "Tank1_Vlv":P;

   // TANK 2 DISCHARGE VALVE
         L     "Var_System_DB".Tk102.Vlv_Actuator_Cmd;
         T     "Tank2_Vlv":P;

   // TANK 3 DISCHARGE VALVE
         L     "Var_System_DB".Tk103.Vlv_Actuator_Cmd;
         T     "Tank3_Vlv":P;

   // SIRUPE VALVE
         L     "Var_System_DB".Sirupe_Valve.Vlv_Actuator_Cmd;
         T     "Sirupe_Vlv":P;

   // WATER VALVE
         L     "Var_System_DB".Water_Valve.Vlv_Actuator_Cmd;
         T     "Water_Vlv":P;

   // MIXER VF
         L     "Var_System_DB".Mixer_Motor.PV;
         T     "Motor_VF":P;
END_REGION

REGION Network 2: *****************************VALVE ACTUATORS********************************************/
   // TANK 1 DISCHARGE AND FILLING VALVES
         A     "Man_Dis_Tk1_Vlv";
         JCN   _001;
         L     27648;
         T     "Var_System_DB".Tk101.Vlv_Actuator_Cmd;
   _001: NOP   0;

         A     "Var_System_DB".TK101_FILLING_VLV.Open_Vlv_Cmd;
         =     "Filling_Vlv1";

   // TANK 2 DISCHARGE AND FILLING VALVES
         A     "Var_System_DB".Tk102.Vlv_Open_Cmd;
         =     "Discharge_Vlv2";

         A     "Var_System_DB".TK102_FILLING_VLV.Open_Vlv_Cmd;
         =     "Filling_Vlv2";

   // TANK 3 DISCHARGE AND FILLING VALVES
         A     "Var_System_DB".Tk103.Vlv_Open_Cmd;
         =     "Discharge_Vlv3";

         A     "Var_System_DB".TK103_FILLING_VLV.Open_Vlv_Cmd;
         =     "Filling_Vlv3";

   // SCALE VALVE
         A     "Var_System_DB".Scale_Discharge_Vlv.Open_Vlv;
         O     "HMI_VAR".Man_Valves.Scale_Vlv;
         =     "Scale_Dis_Vlv";
END_REGION
